// TIA Portal project "Project2_Pompe" (V15.1)

(* hardware
DEVICE "S71500/ET200MP station_1"  S7-1500 station
   slot 0: "Rail_0"  Rack  6ES7 590-1***0-0AA0
   slot 1: "PLC_1"  CPU 1513-1 PN  6ES7 513-1AL02-0AB0  V2.6
      slot 3: "CPU display_1"  6ES7591-1AA00-0AA0
DEVICE "HMI_1"  KTP900 Basic PN
   slot 0: "HMI_1"  KTP900 Basic PN  6AV2 123-2JB03-0AX0  15.1.0.0
   slot 1: "HMI_RT_1"  KTP900 Basic PN  6AV2 123-2JB03-0AX0  15.1.0.0
   slot 5: "HMI_1.IE_CP_1"  PROFINET Interface  15.0.1.0
      slot 1: "PROFINET Interface_1"  PROFINET Interface
         slot 1: "Port_1"  Port
*)

// ===== PLC "PLC_1"  CPU 1513-1 PN =====

VAR_GLOBAL   // PLC tag table "Default tag table"
   "Clock_Byte" AT %MB0 : Byte;
   "Clock_10Hz" AT %M0.0 : Bool;
   "Clock_5Hz" AT %M0.1 : Bool;
   "Clock_2.5Hz" AT %M0.2 : Bool;
   "Clock_2Hz" AT %M0.3 : Bool;
   "Clock_1.25Hz" AT %M0.4 : Bool;
   "Clock_1Hz" AT %M0.5 : Bool;
   "Clock_0.625Hz" AT %M0.6 : Bool;
   "Clock_0.5Hz" AT %M0.7 : Bool;
END_VAR

VAR_GLOBAL   // PLC tag table "Motor1"
   "permisie_start_1" AT %I0.0 : Bool;
   "motor_pornit_1" AT %I0.1 : Bool;
   "temporizare_k4_1" AT %I0.2 : Bool;
   "urgenta_bit_1" AT %I0.4 : Bool;
   "s1_1" AT %I0.7 : Bool;
   "s2_1" AT %I1.0 : Bool;
   "stop1" AT %I1.1 : Bool;
   "ptc1" AT %I1.2 : Bool;
   "timp_oprire_1" AT %ID1 : Time;
   "k1_1" AT %I1.4 : Bool;
   "k2_1" AT %I1.5 : Bool;
   "k3_1" AT %I1.6 : Bool;
   "k4_1" AT %I1.7 : Bool;
   "reset_urgenta_1" AT %I7.0 : Bool;
   "et_k4_1" AT %ID11 : Time;
   "et_stop_1" AT %ID10 : Time;
   "inactiv_1" AT %ID20 : Time;
END_VAR

VAR_GLOBAL   // PLC tag table "Motor2"
   "permisie_start_2" AT %I2.0 : Bool;
   "motor_pornit_2" AT %I2.1 : Bool;
   "temporizare_k4_2" AT %I2.2 : Bool;
   "urgenta_bit_2" AT %I2.3 : Bool;
   "s1_2" AT %I2.4 : Bool;
   "s2_2" AT %I2.5 : Bool;
   "stop2" AT %I2.6 : Bool;
   "ptc2" AT %I2.7 : Bool;
   "timp_oprire_2" AT %ID3 : Time;
   "k1_2" AT %I3.1 : Bool;
   "k2_2" AT %I3.2 : Bool;
   "k3_2" AT %I3.3 : Bool;
   "k4_2" AT %I3.4 : Bool;
   "reset_urgenta_2" AT %I7.1 : Bool;
   "et_k4_2" AT %ID7 : Time;
   "et_stop_2" AT %ID12 : Time;
   "inactiv_2" AT %ID16 : Time;
END_VAR

VAR_GLOBAL   // PLC tag table "Ambele_motoare"
   "ss" AT %I0.6 : Bool;
END_VAR

DATA_BLOCK "db_time"   // DB1
{ S7_Optimized_Access := 'TRUE' }
VERSION : 0.1
   VAR
      timp_inactiv_1 : Time := T#5s;
      timp_inactiv_2 : Time := T#5s;
      timp_et_k4_1 : Time;
      timp_et_k4_2 : Time;
      timp_et_stop_1 : Time;
      timp_et_stop_2 : Time;
      timp_force_sd : Time;
   END_VAR
BEGIN
END_DATA_BLOCK

DATA_BLOCK "db_timp_secunde"   // DB2
{ S7_Optimized_Access := 'TRUE' }
VERSION : 0.1
   VAR
      timp_inactiv_1s : Time := T#5s;
      timp_inactiv_2s : Time := T#5s;
      timp_et_k4_1s : Time;
      timp_et_k4_2s : Time;
      timp_et_stop_1s : Time;
      timp_et_stop_2s : Time;
      timp_sd_secunde : Time;
   END_VAR
BEGIN
END_DATA_BLOCK

DATA_BLOCK "Motor1"   // DB3
{ S7_Optimized_Access := 'TRUE' }
VERSION : 0.1
// stored: InstanceOfName Fct_Motor
"Fct_Motor"
BEGIN
END_DATA_BLOCK

DATA_BLOCK "Motor2"   // DB4
{ S7_Optimized_Access := 'TRUE' }
VERSION : 0.1
// stored: InstanceOfName Fct_Motor
"Fct_Motor"
BEGIN
END_DATA_BLOCK

DATA_BLOCK "db_timp_trecut"   // DB5
{ S7_Optimized_Access := 'TRUE' }
VERSION : 0.1
   VAR
      trecut_et_k4_1 : Bool;
      trecut_et_k4_2 : Bool;
      trecut_et_stop_1 : Bool;
      trecut_et_stop_2 : Bool;
      trecut_inactiv_1 : Bool;
      trecut_inactiv_2 : Bool;
   END_VAR
BEGIN
END_DATA_BLOCK

// folder: System blocks/Program resources

DATA_BLOCK "IEC_Timer_0_DB"   // DB6
{ S7_Optimized_Access := 'TRUE' }
AUTHOR : Simatic
FAMILY : IEC
NAME : IEC_TMR
VERSION : 1.0
// stored: InstanceOfName IEC_TIMER
"IEC_TIMER"
BEGIN
END_DATA_BLOCK

DATA_BLOCK "IEC_Timer_0_DB_1"   // DB7
{ S7_Optimized_Access := 'TRUE' }
AUTHOR : Simatic
FAMILY : IEC
NAME : IEC_TMR
VERSION : 1.0
// stored: InstanceOfName IEC_TIMER
"IEC_TIMER"
BEGIN
END_DATA_BLOCK

// folder: (top level)

FUNCTION_BLOCK "Fct_Motor"   // FB1, LAD
{ S7_Optimized_Access := 'TRUE' }
VERSION : 0.1
   VAR_OUTPUT
      k1 : Bool;
      k2 : Bool;
      k3 : Bool;
      k4 : Bool;
   END_VAR
   VAR_IN_OUT
      "permisie start" : Bool;
      "motor pornit" : Bool;
      "temporizare k4" : Bool;
      "reset urgenta" : Bool;
      "urgenta bit" : Bool;
      s1 : Bool;
      s2 : Bool;
      ss : Bool;
      stop : Bool;
      ptc : Bool;
      et_stop : Time := T#0s;
      et_k4 : Time := T#0s;
      timp_inactiv : Time := T#0s;
   END_VAR
   VAR
      timerK4 : TON_TIME;
      timer_stop : TON_TIME;
   END_VAR
BEGIN

REGION Network 1: selecteaza k1
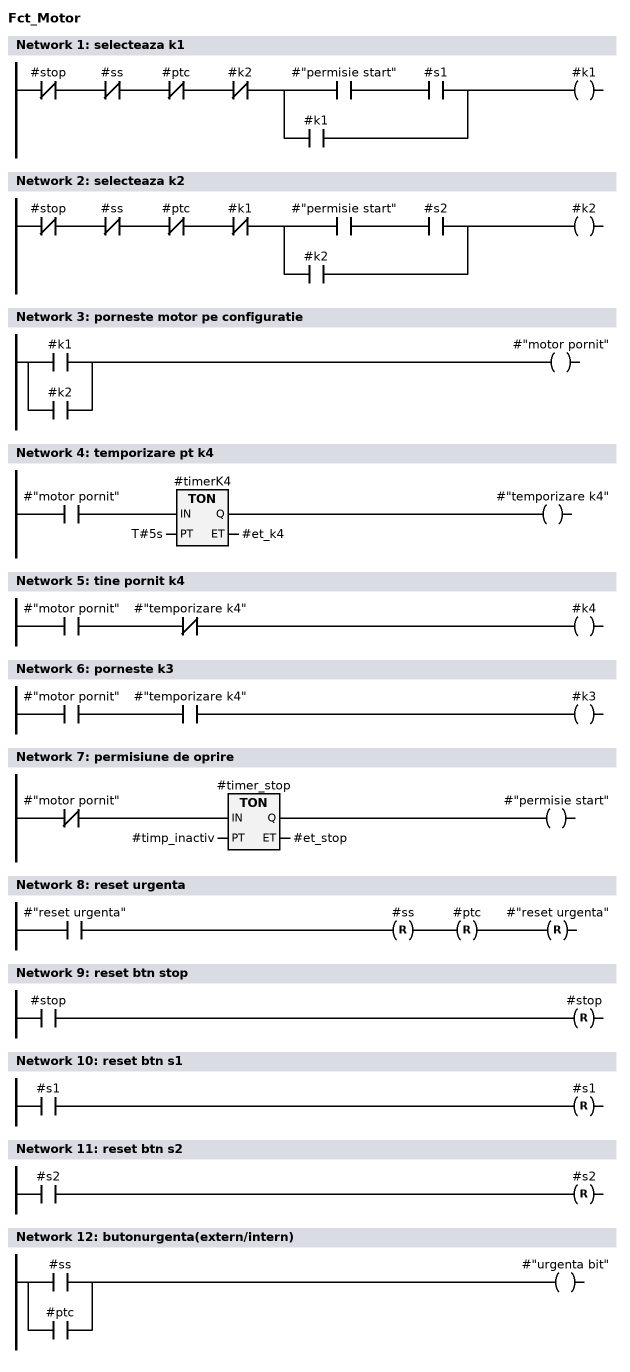
   RUNG wire#powerrail
      I_Contact( #stop )
      I_Contact( #ss )
      I_Contact( #ptc )
      I_Contact( #k2 )
      wire#w1
      Contact( #"permisie start" )
      Contact( #s1 )
      wire#w2
      Coil( #k1 )
   END_RUNG
   RUNG wire#w1
      Contact( #k1 )
   END_RUNG wire#w2
   // the same network as SCL:
   #k1 := NOT #stop AND NOT #ss AND NOT #ptc AND NOT #k2 AND ((#"permisie start" AND #s1) OR #k1);
END_REGION

REGION Network 2: selecteaza k2
   RUNG wire#powerrail
      I_Contact( #stop )
      I_Contact( #ss )
      I_Contact( #ptc )
      I_Contact( #k1 )
      wire#w1
      Contact( #"permisie start" )
      Contact( #s2 )
      wire#w2
      Coil( #k2 )
   END_RUNG
   RUNG wire#w1
      Contact( #k2 )
   END_RUNG wire#w2
   // the same network as SCL:
   #k2 := NOT #stop AND NOT #ss AND NOT #ptc AND NOT #k1 AND ((#"permisie start" AND #s2) OR #k2);
END_REGION

REGION Network 3: porneste motor pe configuratie
   RUNG wire#powerrail
      Contact( #k1 )
      wire#w1
      Coil( #"motor pornit" )
   END_RUNG
   RUNG wire#powerrail
      Contact( #k2 )
   END_RUNG wire#w1
   // the same network as SCL:
   #"motor pornit" := #k1 OR #k2;
END_REGION

REGION Network 4: temporizare pt k4
   #timerK4(IN := #"motor pornit", PT := T#5s, ET => #et_k4);   // TON
   #"temporizare k4" := #timerK4.Q;
END_REGION

REGION Network 5: tine pornit k4
   RUNG wire#powerrail
      Contact( #"motor pornit" )
      I_Contact( #"temporizare k4" )
      Coil( #k4 )
   END_RUNG
   // the same network as SCL:
   #k4 := #"motor pornit" AND NOT #"temporizare k4";
END_REGION

REGION Network 6: porneste k3
   RUNG wire#powerrail
      Contact( #"motor pornit" )
      Contact( #"temporizare k4" )
      Coil( #k3 )
   END_RUNG
   // the same network as SCL:
   #k3 := #"motor pornit" AND #"temporizare k4";
END_REGION

REGION Network 7: permisiune de oprire
   #timer_stop(IN := NOT #"motor pornit", PT := #timp_inactiv, ET => #et_stop);   // TON
   #"permisie start" := #timer_stop.Q;
END_REGION

REGION Network 8: reset urgenta
   RUNG wire#powerrail
      Contact( #"reset urgenta" )
      R_Coil( #ss )
      R_Coil( #ptc )
      R_Coil( #"reset urgenta" )
   END_RUNG
   // the same network as SCL:
   IF #"reset urgenta" THEN
       #ss := FALSE;
       #ptc := FALSE;
       #"reset urgenta" := FALSE;
   END_IF;
END_REGION

REGION Network 9: reset btn stop
   RUNG wire#powerrail
      Contact( #stop )
      R_Coil( #stop )
   END_RUNG
   // the same network as SCL:
   IF #stop THEN #stop := FALSE; END_IF;
END_REGION

REGION Network 10: reset btn s1
   RUNG wire#powerrail
      Contact( #s1 )
      R_Coil( #s1 )
   END_RUNG
   // the same network as SCL:
   IF #s1 THEN #s1 := FALSE; END_IF;
END_REGION

REGION Network 11: reset btn s2
   RUNG wire#powerrail
      Contact( #s2 )
      R_Coil( #s2 )
   END_RUNG
   // the same network as SCL:
   IF #s2 THEN #s2 := FALSE; END_IF;
END_REGION

REGION Network 12: butonurgenta(extern/intern)
   RUNG wire#powerrail
      Contact( #ss )
      wire#w1
      Coil( #"urgenta bit" )
   END_RUNG
   RUNG wire#powerrail
      Contact( #ptc )
   END_RUNG wire#w1
   // the same network as SCL:
   #"urgenta bit" := #ss OR #ptc;
END_REGION
END_FUNCTION_BLOCK

ORGANIZATION_BLOCK "Main"   // OB1, LAD, ProgramCycle
TITLE = "Main Program Sweep (Cycle)"
{ S7_Optimized_Access := 'TRUE' }
VERSION : 0.1
   VAR_INPUT
      Initial_Call : Bool;   // Initial call of this OB
      Remanence : Bool;   // =True, if remanent data are available
   END_VAR
   VAR_TEMP   // added for the SCL form of the ladder/FBD networks
      _w1 : Bool;
   END_VAR
BEGIN

REGION Network 1: initializam motoarele
   // ramas de adaugat sa se vada timerele(partea de ms to s) si sa poti schimba timpul cat e oprit motorul
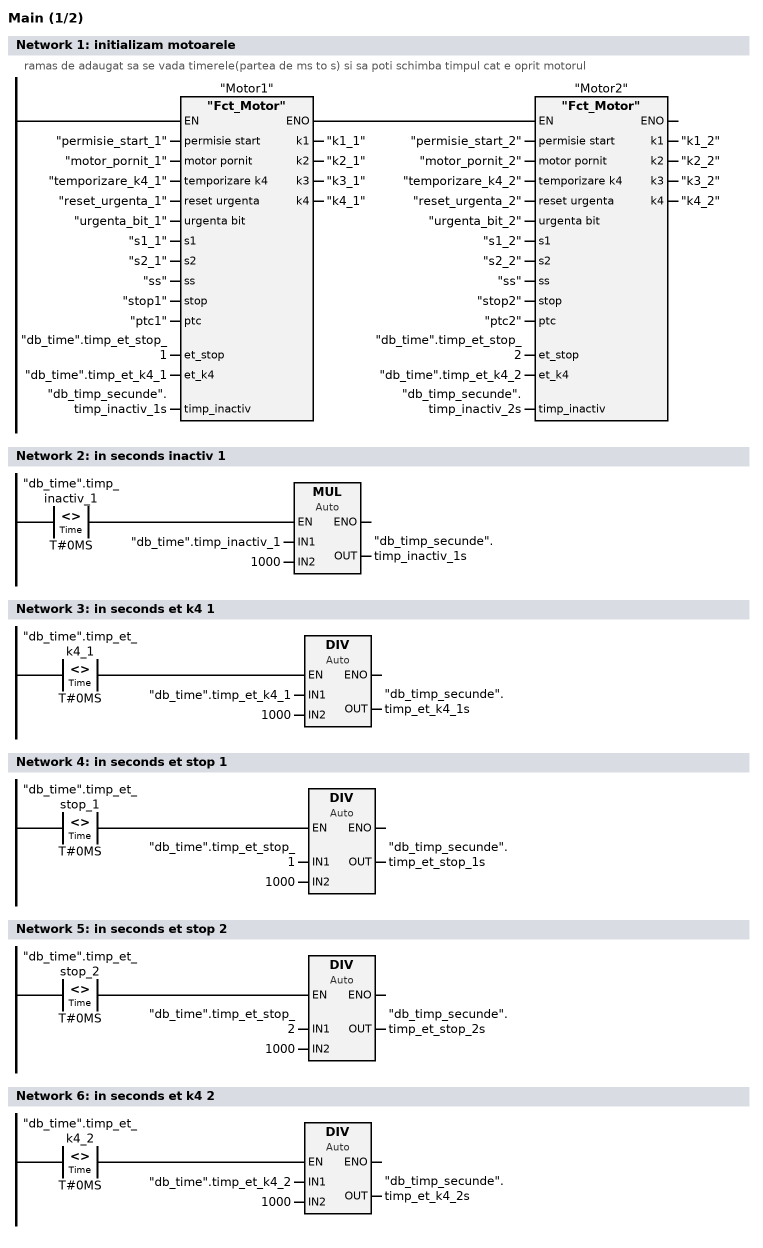
   RUNG wire#powerrail
      "Motor1"("permisie start" := "permisie_start_1", "motor pornit" := "motor_pornit_1", "temporizare k4" := "temporizare_k4_1", "reset urgenta" := "reset_urgenta_1", "urgenta bit" := "urgenta_bit_1", s1 := "s1_1", s2 := "s2_1", ss := "ss", stop := "stop1", ptc := "ptc1", et_stop := "db_time".timp_et_stop_1, et_k4 := "db_time".timp_et_k4_1, timp_inactiv := "db_timp_secunde".timp_inactiv_1s, k1 => "k1_1", k2 => "k2_1", k3 => "k3_1", k4 => "k4_1")
      "Motor2"("permisie start" := "permisie_start_2", "motor pornit" := "motor_pornit_2", "temporizare k4" := "temporizare_k4_2", "reset urgenta" := "reset_urgenta_2", "urgenta bit" := "urgenta_bit_2", s1 := "s1_2", s2 := "s2_2", ss := "ss", stop := "stop2", ptc := "ptc2", et_stop := "db_time".timp_et_stop_2, et_k4 := "db_time".timp_et_k4_2, timp_inactiv := "db_timp_secunde".timp_inactiv_2s, k1 => "k1_2", k2 => "k2_2", k3 => "k3_2", k4 => "k4_2")
   END_RUNG
   // the same network as SCL:
   "Motor1"("permisie start" := "permisie_start_1",   // "Fct_Motor"
            "motor pornit" := "motor_pornit_1",
            "temporizare k4" := "temporizare_k4_1",
            "reset urgenta" := "reset_urgenta_1",
            "urgenta bit" := "urgenta_bit_1",
            s1 := "s1_1",
            s2 := "s2_1",
            ss := "ss",
            stop := "stop1",
            ptc := "ptc1",
            et_stop := "db_time".timp_et_stop_1,
            et_k4 := "db_time".timp_et_k4_1,
            timp_inactiv := "db_timp_secunde".timp_inactiv_1s,
            k1 => "k1_1",
            k2 => "k2_1",
            k3 => "k3_1",
            k4 => "k4_1",
            ENO => #_w1);
   IF #_w1 THEN
       "Motor2"("permisie start" := "permisie_start_2",   // "Fct_Motor"
                "motor pornit" := "motor_pornit_2",
                "temporizare k4" := "temporizare_k4_2",
                "reset urgenta" := "reset_urgenta_2",
                "urgenta bit" := "urgenta_bit_2",
                s1 := "s1_2",
                s2 := "s2_2",
                ss := "ss",
                stop := "stop2",
                ptc := "ptc2",
                et_stop := "db_time".timp_et_stop_2,
                et_k4 := "db_time".timp_et_k4_2,
                timp_inactiv := "db_timp_secunde".timp_inactiv_2s,
                k1 => "k1_2",
                k2 => "k2_2",
                k3 => "k3_2",
                k4 => "k4_2");
   END_IF;
END_REGION

REGION Network 2: in seconds inactiv 1
   RUNG wire#powerrail
      { S7_Templates := "SrcType := Time" } NE_Contact(in1 := "db_time".timp_inactiv_1, in2 := T#0MS)
      Mul(in1 := "db_time".timp_inactiv_1, in2 := 1000, out => "db_timp_secunde".timp_inactiv_1s)
   END_RUNG
   // the same network as SCL:
   IF "db_time".timp_inactiv_1 <> T#0MS THEN
       "db_timp_secunde".timp_inactiv_1s := "db_time".timp_inactiv_1 * 1000;
   END_IF;
END_REGION

REGION Network 3: in seconds et k4 1
   RUNG wire#powerrail
      { S7_Templates := "SrcType := Time" } NE_Contact(in1 := "db_time".timp_et_k4_1, in2 := T#0MS)
      Div(in1 := "db_time".timp_et_k4_1, in2 := 1000, out => "db_timp_secunde".timp_et_k4_1s)
   END_RUNG
   // the same network as SCL:
   IF "db_time".timp_et_k4_1 <> T#0MS THEN
       "db_timp_secunde".timp_et_k4_1s := "db_time".timp_et_k4_1 / 1000;
   END_IF;
END_REGION

REGION Network 4: in seconds et stop 1
   RUNG wire#powerrail
      { S7_Templates := "SrcType := Time" } NE_Contact(in1 := "db_time".timp_et_stop_1, in2 := T#0MS)
      Div(in1 := "db_time".timp_et_stop_1, in2 := 1000, out => "db_timp_secunde".timp_et_stop_1s)
   END_RUNG
   // the same network as SCL:
   IF "db_time".timp_et_stop_1 <> T#0MS THEN
       "db_timp_secunde".timp_et_stop_1s := "db_time".timp_et_stop_1 / 1000;
   END_IF;
END_REGION

REGION Network 5: in seconds et stop 2
   RUNG wire#powerrail
      { S7_Templates := "SrcType := Time" } NE_Contact(in1 := "db_time".timp_et_stop_2, in2 := T#0MS)
      Div(in1 := "db_time".timp_et_stop_2, in2 := 1000, out => "db_timp_secunde".timp_et_stop_2s)
   END_RUNG
   // the same network as SCL:
   IF "db_time".timp_et_stop_2 <> T#0MS THEN
       "db_timp_secunde".timp_et_stop_2s := "db_time".timp_et_stop_2 / 1000;
   END_IF;
END_REGION

REGION Network 6: in seconds et k4 2
   RUNG wire#powerrail
      { S7_Templates := "SrcType := Time" } NE_Contact(in1 := "db_time".timp_et_k4_2, in2 := T#0MS)
      Div(in1 := "db_time".timp_et_k4_2, in2 := 1000, out => "db_timp_secunde".timp_et_k4_2s)
   END_RUNG
   // the same network as SCL:
   IF "db_time".timp_et_k4_2 <> T#0MS THEN
       "db_timp_secunde".timp_et_k4_2s := "db_time".timp_et_k4_2 / 1000;
   END_IF;
END_REGION

REGION Network 7: in seconds incativ 2
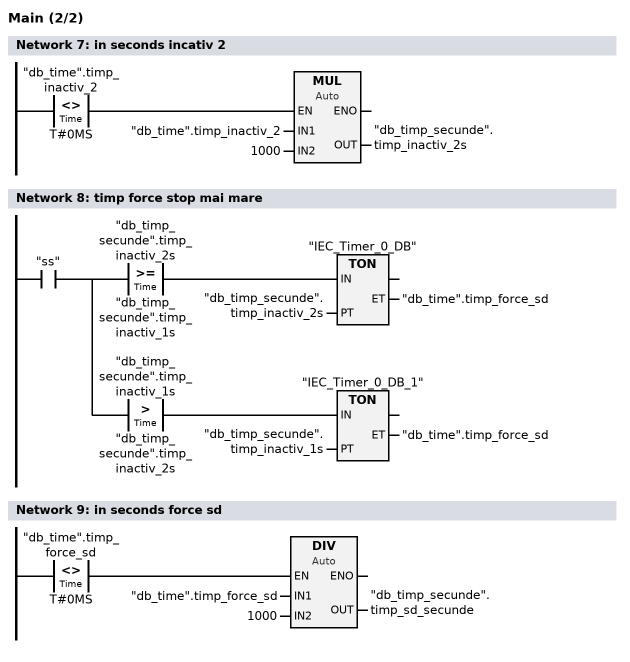
   RUNG wire#powerrail
      { S7_Templates := "SrcType := Time" } NE_Contact(in1 := "db_time".timp_inactiv_2, in2 := T#0MS)
      Mul(in1 := "db_time".timp_inactiv_2, in2 := 1000, out => "db_timp_secunde".timp_inactiv_2s)
   END_RUNG
   // the same network as SCL:
   IF "db_time".timp_inactiv_2 <> T#0MS THEN
       "db_timp_secunde".timp_inactiv_2s := "db_time".timp_inactiv_2 * 1000;
   END_IF;
END_REGION

REGION Network 8: timp force stop mai mare
   "IEC_Timer_0_DB".TON(IN := "ss" AND ("db_timp_secunde".timp_inactiv_2s >= "db_timp_secunde".timp_inactiv_1s),
                        PT := "db_timp_secunde".timp_inactiv_2s,
                        ET => "db_time".timp_force_sd);
   "IEC_Timer_0_DB_1".TON(IN := "ss" AND ("db_timp_secunde".timp_inactiv_1s > "db_timp_secunde".timp_inactiv_2s),
                          PT := "db_timp_secunde".timp_inactiv_1s,
                          ET => "db_time".timp_force_sd);
END_REGION

REGION Network 9: in seconds force sd
   RUNG wire#powerrail
      { S7_Templates := "SrcType := Time" } NE_Contact(in1 := "db_time".timp_force_sd, in2 := T#0MS)
      Div(in1 := "db_time".timp_force_sd, in2 := 1000, out => "db_timp_secunde".timp_sd_secunde)
   END_RUNG
   // the same network as SCL:
   IF "db_time".timp_force_sd <> T#0MS THEN
       "db_timp_secunde".timp_sd_secunde := "db_time".timp_force_sd / 1000;
   END_IF;
END_REGION
END_ORGANIZATION_BLOCK

(* ===== HMI "HMI_RT_1" =====
system functions are stored by id; their names below are inferred from use
connection "HMI_Connection_1": ETHERNET, SMART_S7_1500_OMS

HMI tags "Default tag table"
   "stop1" : Bool = PLC stop1 AT %I1.1, 1 s
   "s1_1" : Bool = PLC s1_1 AT %I0.7, 1 s
   "s2_1" : Bool = PLC s2_1 AT %I1.0, 1 s
   "k1_1" : Bool = PLC k1_1 AT %I1.4, 1 s
   "k2_1" : Bool = PLC k2_1 AT %I1.5, 1 s
   "urgenta_bit_1" : Bool = PLC urgenta_bit_1 AT %I0.4, 1 s
   "ptc1" : Bool = PLC ptc1 AT %I1.2, 1 s
   "k4_1" : Bool = PLC k4_1 AT %I1.7, 1 s
   "k3_1" : Bool = PLC k3_1 AT %I1.6, 1 s
   "timp_oprire_1" : Time = PLC timp_oprire_1 AT %ID1, 1 s
   "motor_pornit_1" : Bool = PLC motor_pornit_1 AT %I0.1, 1 s
   "stop2" : Bool = PLC stop2 AT %I2.6, 1 s
   "s1_2" : Bool = PLC s1_2 AT %I2.4, 1 s
   "s2_2" : Bool = PLC s2_2 AT %I2.5, 1 s
   "k1_2" : Bool = PLC k1_2 AT %I3.1, 1 s
   "k2_2" : Bool = PLC k2_2 AT %I3.2, 1 s
   "urgenta_bit_2" : Bool = PLC urgenta_bit_2 AT %I2.3, 1 s
   "ptc2" : Bool = PLC ptc2 AT %I2.7, 1 s
   "reset_urgenta_1" : Bool = PLC reset_urgenta_1 AT %I7.0, 1 s
   "reset_urgenta_2" : Bool = PLC reset_urgenta_2 AT %I7.1, 1 s
   "k4_2" : Bool = PLC k4_2 AT %I3.4, 1 s
   "k3_2" : Bool = PLC k3_2 AT %I3.3, 1 s
   "motor_pornit_2" : Bool = PLC motor_pornit_2 AT %I2.1, 1 s
   "ss" : Bool = PLC ss AT %I0.6, 1 s
   "et_k4_1" : Time = PLC et_k4_1 AT %ID11, 1 s
   "et_stop_1" : Time = PLC et_stop_1 AT %ID10, 1 s
   "et_stop_2" : Time = PLC et_stop_2 AT %ID12, 1 s
   "et_k4_2" : Time = PLC et_k4_2 AT %ID7, 1 s
   "inactiv_2" : Time = PLC inactiv_2 AT %ID16, 1 s
   "inactiv_1" : Time = PLC inactiv_1 AT %ID20, 1 s
   "db_time_timp_et_stop_1" : Time = PLC db_time.timp_et_stop_1, 1 s
   "db_time_timp_et_k4_1" : Time = PLC db_time.timp_et_k4_1, 1 s
   "db_time_timp_inactiv_1" : Time = PLC db_time.timp_inactiv_1, 1 s
   "db_time_timp_et_stop_2" : Time = PLC db_time.timp_et_stop_2, 1 s
   "db_time_timp_inactiv_2" : Time = PLC db_time.timp_inactiv_2, 1 s
   "db_time_timp_et_k4_2" : Time = PLC db_time.timp_et_k4_2, 1 s
   "db_time_timp_force_sd" : Time = PLC db_time.timp_force_sd, 1 s
   "db_timp_secunde_timp_et_stop_1s" : Time = PLC db_timp_secunde.timp_et_stop_1s, 1 s
   "db_timp_secunde_timp_inactiv_1s" : Time = PLC db_timp_secunde.timp_inactiv_1s, 1 s
   "db_timp_secunde_timp_et_k4_1s" : Time = PLC db_timp_secunde.timp_et_k4_1s, 1 s
   "db_timp_secunde_timp_et_stop_2s" : Time = PLC db_timp_secunde.timp_et_stop_2s, 1 s
   "db_timp_secunde_timp_inactiv_2s" : Time = PLC db_timp_secunde.timp_inactiv_2s, 1 s
   "db_timp_secunde_timp_et_k4_2s" : Time = PLC db_timp_secunde.timp_et_k4_2s, 1 s
   "db_timp_secunde_timp_sd_secunde" : Time = PLC db_timp_secunde.timp_sd_secunde, 1 s

Template "Template_1" 800x480
   Button "Exit" at 722,440 size 55x39; TextOff 'Exit'; PictureOff "ExitRuntime_KTP900_Basic_PN_TR"; PictureOn "ExitRuntime_KTP900_Basic_PN_TR"
      on Release: StopRuntime(0)
   Button "Template_Button" at 622,440 size 55x39; TextOff 'Text'
   Button "Template_Button_1" at 522,440 size 55x39; TextOff 'Text'
   Button "Template_Button_2" at 422,440 size 55x39; TextOff 'Text'
   Button "Template_Button_3" at 322,440 size 55x39; TextOff 'Text'
   Button "Template_Button_4" at 222,440 size 55x39; TextOff 'Text'
   Button "Alarms" at 122,440 size 55x39; TextOff 'Alarms'; PictureOff "AlarmDisplay_KTP900_Basic_PN_TR"; PictureOn "AlarmDisplay_KTP900_Basic_PN_TR"
      on Release: function_ef3f5d25("Alarm window_Unacknowledged", -1)
   Button "Start screen" at 22,440 size 55x39; TextOff 'Start screen'; PictureOff "NavigateHome_KTP900_Basic_PN_TR"; PictureOn "NavigateHome_KTP900_Basic_PN_TR"
      on Release: ActivateScreen("Root screen", 0)
   DateTimeField "HmiScreenItemData" at 695,20 size 105x20
   DateTimeField "HmiScreenItemData_1" at 695,0 size 105x20
   GraphicView "Logo" at 0,0 size 71x40; Picture "Logo of HMI_1"

screen "Root screen" 800x480, template "Template_1"
   Circle "Circle_1" at 129,113 size 86x86
      Appearance <- "motor_pornit_1"
   Group "Group" at 129,113 size 89x87
   TextField "Text field_1" at 156,61 size 35x20; Text 'Stop'
   TextField "Text field_2" at 18,64 size 67x20; Text 'Clockwise'
   TextField "Text field_3" at 256,66 size 87x20; Text 'CtrClockwise'
   Button "Button_1" at 657,68 size 96x32; TextOff 'Stop'
      on Click: SetBit("stop1")
   TextField "Text field_4" at 619,73 size 21x20; Text 'S0'
   Button "Button_2" at 658,118 size 96x32; TextOff 'Start K1'
      on Click: SetBit("s1_1")
   Button "Button_3" at 658,167 size 96x32; TextOff 'Start K2'
      on Click: SetBit("s2_1")
   Circle "Circle_3" at 606,113 size 42x42
      Appearance <- "k1_1"
   Circle "Circle_4" at 606,168 size 42x42
      Appearance <- "k2_1"
   TextField "Text field_5" at 570,122 size 21x20; Text 'S1'
   TextField "Text field_6" at 570,175 size 21x20; Text 'S2'
   Button "Button_4" at 623,351 size 96x32; TextOff 'ESD'
      on Click: SetBit("ptc1")
   TextField "Text field_7" at 584,353 size 21x20; Text 'SS'
   Circle "Circle_2" at 331,307 size 79x79
      Appearance <- "k3_1"
   Circle "Circle_5" at 440,306 size 79x79
      Appearance <- "k4_1"
   TextField "Text field_8" at 362,334 size 21x20; Text 'K3'
   TextField "Text field_9" at 473,336 size 21x20; Text 'K4'
   Button "Button_5" at 21,390 size 96x32; TextOff 'Just press'
   Button "Button_6" at 623,397 size 96x32; TextOff 'Reset ESD'
      on Click: SetBit("reset_urgenta_1")
   Circle "Circle_6" at 128,271 size 101x101
      Appearance <- "motor_pornit_1"
   TextField "Text field_12" at 73,307 size 44x20; Text 'Motor'
   Group "Group_1" at 262,108 size 89x87
   Group "Group_2" at 17,114 size 89x87
   Ellipse "Ellipse_1" at 640,317 size 67x28
      Appearance <- "urgenta_bit_1"
   TextField "Text field_13" at 378,16 size 56x20; Text 'Motor 1'
   Button "Button_7" at 681,263 size 96x32; TextOff 'Next'
      on Click: ActivateScreen("Screen_1", 0)
   IOField "I/O field_1" at 438,265 size 96x32; FormatPattern 9999; Unit s
      ProcessValue <- "db_timp_secunde_timp_et_k4_1s"
   TextField "Text field_10" at 446,228 size 53x20; Text 'Time k4'
   IOField "I/O field_2" at 510,61 size 96x32; FormatPattern 9999; Unit s
      ProcessValue <- "db_timp_secunde_timp_et_stop_1s"
   TextField "Text field_11" at 536,36 size 73x20; Text 'Timer stop'
   IOField "I/O field_3" at 437,165 size 96x32; FormatPattern 99; Unit s
      ProcessValue <- "db_time_timp_inactiv_1"
   TextField "Text field_14" at 421,136 size 114x20; Text 'Set time inactive'
   Circle "Circle_7" at 262,108 size 86x86
      Appearance <- "k2_1"
   Circle "Circle_8" at 17,114 size 86x86
      Appearance <- "k1_1"

screen "Screen_1" 800x480
   Circle "Circle_1" at 129,113 size 86x86
      Appearance <- "motor_pornit_2"
   Group "Group" at 129,113 size 89x87
   TextField "Text field_1" at 156,61 size 35x20; Text 'Stop'
   TextField "Text field_2" at 18,64 size 67x20; Text 'Clockwise'
   TextField "Text field_3" at 256,66 size 87x20; Text 'CtrClockwise'
   Button "Button_1" at 657,68 size 96x32; TextOff 'Stop'
      on Click: SetBit("stop2")
   TextField "Text field_4" at 619,73 size 21x20; Text 'S0'
   Button "Button_2" at 658,118 size 96x32; TextOff 'Start K1'
      on Click: SetBit("s1_2")
   Button "Button_3" at 658,167 size 96x32; TextOff 'Start K2'
      on Click: SetBit("s2_2")
   Circle "Circle_3" at 606,113 size 42x42
      Appearance <- "k1_2"
   Circle "Circle_4" at 606,168 size 42x42
      Appearance <- "k2_2"
   TextField "Text field_5" at 570,122 size 21x20; Text 'S1'
   TextField "Text field_6" at 570,175 size 21x20; Text 'S2'
   Button "Button_4" at 623,351 size 96x32; TextOff 'ESD'
      on Click: SetBit("ptc2")
   TextField "Text field_7" at 584,353 size 21x20; Text 'SS'
   Circle "Circle_2" at 331,307 size 79x79
      Appearance <- "k3_2"
   Circle "Circle_5" at 440,306 size 79x79
      Appearance <- "k4_2"
   TextField "Text field_8" at 362,334 size 21x20; Text 'K3'
   TextField "Text field_9" at 473,336 size 21x20; Text 'K4'
   Button "Button_5" at 21,390 size 96x32; TextOff 'Just press'
   Button "Button_6" at 623,397 size 96x32; TextOff 'Reset ESD'
      on Click: SetBit("reset_urgenta_2")
   Circle "Circle_6" at 128,271 size 101x101
      Appearance <- "motor_pornit_2"
   TextField "Text field_12" at 73,307 size 44x20; Text 'Motor'
   Group "Group_1" at 262,108 size 89x87
   Group "Group_2" at 17,114 size 89x87
   Ellipse "Ellipse_1" at 640,317 size 67x28
      Appearance <- "urgenta_bit_2"
   TextField "Text field_13" at 375,9 size 52x20; Text 'Motor2'
   Button "Button_7" at 699,255 size 96x32; TextOff 'Next'
      on Click: ActivateScreen("Screen_2", 0)
   Button "Button_8" at 599,255 size 96x32; TextOff 'Prev'
      on Click: ActivateScreen("Root screen", 0)
   IOField "I/O field_1" at 438,265 size 96x32; FormatPattern 9999; Unit s
      ProcessValue <- "db_timp_secunde_timp_et_k4_2s"
   IOField "I/O field_2" at 509,58 size 96x32; FormatPattern 9999; Unit s
      ProcessValue <- "db_timp_secunde_timp_et_stop_2s"
   TextField "Text field_10" at 454,237 size 60x20; Text 'Timer K4'
   TextField "Text field_11" at 511,29 size 73x20; Text 'Timer stop'
   IOField "I/O field_3" at 438,157 size 96x32; FormatPattern 99; Unit s
      ProcessValue <- "db_time_timp_inactiv_2"
   TextField "Text field_14" at 427,137 size 114x20; Text 'Set time inactive'
   Circle "Circle_7" at 262,108 size 86x86
      Appearance <- "k2_2"
   Circle "Circle_8" at 17,114 size 86x86
      Appearance <- "k1_2"

screen "Screen_2" 800x480
   Circle "Circle_1" at 115,129 size 79x79
      Appearance <- "motor_pornit_1"
   Circle "Circle_2" at 212,127 size 79x79
      Appearance <- "motor_pornit_2"
   TextField "Text field_1" at 124,95 size 44x20; Text 'M1 on'
   TextField "Text field_2" at 237,96 size 44x20; Text 'M2 on'
   Button "Button_1" at 631,83 size 127x32; TextOff 'Force stop both'
      on Click: SetBit("ss")
   Button "Button_2" at 628,141 size 130x32; TextOff 'Reset force stop'
      on Click: SetBit("reset_urgenta_1"); SetBit("reset_urgenta_2")
   TextField "Text field_3" at 110,279 size 128x20; Text 'M1 going clockwise'
      Visibility <- "k1_1"
   TextField "Text field_4" at 109,308 size 168x20; Text 'M1 going counter clkwise'
      Visibility <- "k2_1"
   TextField "Text field_5" at 379,276 size 113x20; Text 'M2 going clkwise'
      Visibility <- "k1_2"
   TextField "Text field_6" at 379,308 size 172x20; Text 'M2 going counter clkwise'
      Visibility <- "k2_2"
   Button "Button_3" at 656,208 size 96x32; TextOff 'Prev'
      on Click: ActivateScreen("Screen_1", 0)
   Ellipse "Ellipse_1" at 529,37 size 61x37
      Appearance <- "urgenta_bit_1"
   Ellipse "Ellipse_2" at 611,36 size 61x37
      Appearance <- "urgenta_bit_2"
   TextField "Text field_7" at 546,17 size 13x20; Text '1'
   TextField "Text field_8" at 635,13 size 13x20; Text '2'
   IOField "I/O field_1" at 645,308 size 96x32; FormatPattern 9999; Unit s
      ProcessValue <- "db_timp_secunde_timp_sd_secunde"
   TextField "Text field_9" at 648,283 size 77x20; Text 'Stop timer'
*)